// TIA Portal project "CurrentConfig" (V16)

(* hardware
DEVICE "ET 200S station_1"  ET 200S station
   slot 0: "Rack"  Rail
   slot 2: "-20K0 - PLC"  IM151-8 PN/DP CPU  6ES7 151-8AB01-0AB0  V3.2
      slot 1: "PROFINET interface_1"  PN-IO
         slot 1: "Port_1"  Port
         slot 2: "Port_2"  Port
         slot 3: "Port_3"  Port
   slot 4: "-20K1 - VOEDING"  PM-E 24VDC  6ES7 138-4CA01-0AA0
   slot 5: "-20K2 - INGANG_1"  8DI DC24V  6ES7 131-4BF00-0AA0
   slot 6: "-20K3 - INGANG_2"  8DI DC24V  6ES7 131-4BF00-0AA0
   slot 7: "-20K4 - INGANG_3"  8DI DC24V  6ES7 131-4BF00-0AA0
   slot 8: "-20K5 - INGANG_4"  8DI x 24VDC  6ES7 131-4BF00-0AA0
   slot 9: "-20K6 - UITGANG_1"  8DO x 24VDC / 0.5A  6ES7 132-4BF00-0AA0
   slot 10: "8DO x 24VDC / 0.5A_1"  8DO x 24VDC / 0.5A  6ES7 132-4BF00-0AA0
   slot 11: "PM-E 24VDC_1"  PM-E 24VDC  6ES7 138-4CA01-0AA0
   slot 12: "-20K8 - UITGANG_2"  8DO x 24VDC / 0.5A  6ES7 132-4BF00-0AA0
   slot 13: "-20K9 - UITGANG_3"  8DO x 24VDC / 0.5A  6ES7 132-4BF00-0AA0
   slot 14: "-20K10 - UITGANG_4"  8DO x 24VDC / 0.5A  6ES7 132-4BF00-0AA0
   slot 15: "-20K11 - UITGANG_5"  8DO x 24VDC / 0.5A  6ES7 132-4BF00-0AA0
   slot 16: "-20K12 - UITGANG_6 (4)"  4DO x 24VDC / 0.5A ST  6ES7 132-4BD02-0AA0
   slot 17: "-20K13 - UITGANG_7 (4)"  4DO x 24VDC / 0.5A ST  6ES7 132-4BD02-0AA0
   slot 18: "1 Count 24V Encoder Wals"  1 COUNT 24V  6ES7 138-4DA04-0AB0  V2.0
   slot 19: "1 Count 24V Encoder Band"  1 COUNT 24V  6ES7 138-4DA04-0AB0  V2.0
DEVICE "HMI_1"  KTP700 Basic PN
   slot 0: "HMI_1"  KTP700 Basic PN  6AV2 123-2GB03-0AX0  16.0.0.0
   slot 1: "HMI_RT_2"  KTP700 Basic PN  6AV2 123-2GB03-0AX0  16.0.0.0
   slot 5: "HMI_1.IE_CP_1"  PROFINET Interface  16.0.0.0
      slot 1: "PROFINET Interface_1"  PROFINET Interface
         slot 1: "Port_1"  Port
*)

// ===== PLC "-20K0 - PLC"  IM151-8 PN/DP CPU =====

VAR_GLOBAL   // PLC tag table "Default tag table"
   "Drive 1 Ready" AT %I0.0 : Bool;   // +MC-21K2:1 - Drive 1 Ready
   "Drive 2 Ready" AT %I0.1 : Bool;   // +MC-21K2:5 - Drive 2 Ready
   "Drive 3 Ready" AT %I0.2 : Bool;   // +MC-21K2:2 - Drive 3 Ready
   "Drive 4 Ready" AT %I0.3 : Bool;   // +MC-21K2:6 - Drive 4 Ready
   "Drive 5 Ready" AT %I0.4 : Bool;   // +MC-21K2:3 - Drive 5 Ready
   "Sensor Trechter" AT %I0.5 : Bool;   // +MC-21K2:7 - Sensor Trechter
   "Sensor Op Band" AT %I0.6 : Bool;   // +MC-21K2:4 Sensor Op Band
   "Sensor Wals (Option)" AT %I0.7 : Bool;   // +MC-21K2:8 - Sensor Wals (Option)
   "ESB Oke" AT %I1.0 : Bool;   // +MC-21K3:1 - ESB Oke
   "ESB Pressend" AT %I1.1 : Bool;   // +MC-21K3:5 - ESB Pressend
   "Reset Active" AT %I1.2 : Bool;   // +MC-21K3:2 - Reset Active
   "Noodsleutel(1)" AT %I1.3 : Bool;   // +MC-21K3:6 - NOODSLEUTEL
   "Alle uitgangen(1)" AT %I1.4 : Bool;   // +MC-21K3:3 - Alle uitgangen
   "Door 1 NC contact" AT %I1.5 : Bool;   // +MC-21K3:7 - Safety Doorswitch 1
   "Door 1 NO contact" AT %I1.6 : Bool;   // +MC-21K3:4 - Safety Doorswitch 1 Normaly open
   "Door 2 NC contact" AT %I1.7 : Bool;   // +MC-21K3:8 - Safety Doorswitch 2
   "Spare(5)" AT %I3.0 : Bool;
   "Spare(6)" AT %I3.1 : Bool;
   "Spare(10)" AT %I180.0 : Bool;   // Spare
   "Spare(11)" AT %I180.1 : Bool;   // Spare
   "Spare(12)" AT %I3.4 : Bool;   // Spare
   "Spare(13)" AT %I3.5 : Bool;   // Spare
   "Spare(14)" AT %I3.6 : Bool;   // Spare
   "Spare(15)" AT %I3.7 : Bool;   // Spare
   "Programma 1" AT %I2.0 : Bool;   // +MC-21K4:1 - Programma 1
   "Programma 2" AT %I2.1 : Bool;   // +MC-21K4:5 - Programma 2 (Option)
   "Programma 3" AT %I2.2 : Bool;   // +MC-21K4:2 - Programma 3
   "Cleaning" AT %I2.3 : Bool;   // +MC-21K4:6 - Cleaning
   "Start Machine" AT %I2.4 : Bool;   // +MC-21K4:3 - Start Machine
   "Stop Machine" AT %I2.5 : Bool;   // +MC-21K4:7 - Stop Machine
   "Spare(16)" AT %I2.6 : Bool;   // Spare
   "Encoder_Z_Puls" AT %I2.7 : Bool;   // Spare
   "Safety Relais" AT %Q0.0 : Bool;   // +MC-21K6:1 - Safety Relais
   "Bel Storing" AT %Q0.1 : Bool;   // +MC-21K6:5 - Bel Storing
   "Spare" AT %Q5.3 : Bool;   // Spare
   "Drive 1 RUN FWD" AT %Q1.0 : Bool;   // +MC-21K8:1 - Drive 1 RUN FWD
   "Drive 1 REV]" AT %Q1.1 : Bool;   // +MC-21K8:5 - Drive 1 REV
   "Drive 1 Speed 1" AT %Q1.2 : Bool;   // +MC-21K8:2 - Drive 1 Speed 1
   "Drive 1 Speed 2" AT %Q1.3 : Bool;   // +MC-21K8:6 - Drive 1 Speed 2
   "Spare(3)" AT %Q1.4 : Bool;   // Spare
   "Drive 2 RUN FWD" AT %Q1.5 : Bool;   // +MC-21K8:7 - Drive 2 RUN FWD
   "Drive 2 REV" AT %Q1.6 : Bool;   // +MC-21K8:4 - Drive 2 REV
   "Drive 2 Speed 1" AT %Q1.7 : Bool;   // +MC-21K8:8 - Drive 2 Speed 1
   "Drive 2 Speed 2" AT %Q2.0 : Bool;   // +MC-21K9:1 - Drive 2 Speed 2
   "Spare(4)" AT %Q2.1 : Bool;   // Spare
   "Drive 3 RUN FWD" AT %Q2.2 : Bool;   // +MC-21K9:2 - Drive 3 RUN FWD
   "Drive 3 REV" AT %Q2.3 : Bool;   // +MC-21K9:6 - Drive 3 REV
   "Drive 3 Speed 1" AT %Q2.4 : Bool;   // +MC-21K9:3 - Drive 3 Speed 1
   "Drive 3 Speed 2" AT %Q2.5 : Bool;   // +MC-21K9:7 - Drive 3 Speed 2
   "Spare(21)" AT %Q2.6 : Bool;   // Spare
   "Drive 4 RUN FWD" AT %Q2.7 : Bool;   // +MC-21K9:8 - Drive 4 RUN FWD
   "Drive 4 REV" AT %Q3.0 : Bool;   // +MC-21K10:1 - Drive 4 REV
   "Drive 4 Speed 1" AT %Q3.1 : Bool;   // +MC-21K10:5 - Drive 4 Speed 1
   "Drive 4 Speed 2" AT %Q3.2 : Bool;   // +MC-21K10:2 - Drive 4 Speed 2
   "Spare(22)" AT %Q3.3 : Bool;   // Spare
   "Drive 5 RUN FWD" AT %Q3.4 : Bool;   // +MC-21K10:3 - Drive 5 RUN FWD
   "Drive 5 REV" AT %Q3.5 : Bool;   // +MC-21K10:7 - Drive 5 REV
   "Drive 5 Speed 1" AT %Q3.6 : Bool;   // +MC-21K10:4 - Drive 5 Speed 1
   "Drive 5 Speed 2" AT %Q3.7 : Bool;   // +MC-21K10:8 - Drive 5 Speed 2
   "Spare(23)" AT %Q4.0 : Bool;   // Spare
   "LED Programma 1" AT %Q4.1 : Bool;   // +MC-21K11:5 - LED Programma 1
   "LED Programma 2" AT %Q4.2 : Bool;   // +MC-21K11:2 - LED Programma 2
   "LED Programma 3" AT %Q4.3 : Bool;   // +MC-21K11:6 - LED Programma 3
   "LED E-STOP" AT %Q0.2 : Bool;   // +MC-21K6:2- LED E-STOP
   "LED RUN" AT %Q4.5 : Bool;   // +MC-21K11:7 - LED RUN
   "Valve 1" AT %Q4.6 : Bool;   // +MC-21K11:4 - Valve 1
   "Valve 2" AT %Q4.7 : Bool;   // +MC-21K11:8 - Valve 2
   "Valve 3" AT %Q5.0 : Bool;   // +MC-21K12:1 - Valve 3
   "Valve 4" AT %Q5.1 : Bool;   // +MC-21K12:5 - Valve 4
   "Valve 5" AT %Q5.2 : Bool;   // +MC-21K12:2 - Valve 5
   "Spare(1)" AT %Q6.0 : Bool;   // Spare
   "Spare(2)" AT %Q6.1 : Bool;   // Spare
   "Spare(18)" AT %Q6.2 : Bool;   // Spare
   "Spare(19)" AT %Q6.3 : Bool;   // Spare
   "Spare(20)" AT %Q4.4 : Bool;   // Spare
   "Drive 1 Rapid Stop" AT %Q0.3 : Bool;   // +MC-21K6:6 - Drive 1 Rapid Stop
   "Drive 2 Rapid Stop" AT %Q0.4 : Bool;   // +MC-21K6:3 - Drive 2 Rapid Stop
   "Drive 3 Rapid Stop" AT %Q0.5 : Bool;   // +MC-21K6:7 - Drive 3 Rapid Stop
   "Drive 4 Rapid Stop" AT %Q0.6 : Bool;   // +MC-21K6:4 - Drive 4 Rapid Stop
   "Drive 5 Rapid Stop" AT %Q0.7 : Bool;   // +MC-21K6:8 - Drive 5 Rapid Stop
   "Systeem RUN" AT %M0.0 : Bool;   // Systeem RUN
   "Tag_1" AT %M0.1 : Bool;
   "Tag_2" AT %M0.2 : Bool;
   "Tag_3" AT %M0.3 : Bool;
   "Tag_4" AT %M0.4 : Bool;
   "Safety Feedback" AT %M0.6 : Bool;
   "Tag_5" AT %M0.7 : Bool;
   "Tag_6" AT %M1.0 : Bool;
   "ONC Drive 1 RUN FWD" AT %M10.0 : Bool;
   "ONC Drive 2 RUN FWD" AT %M10.1 : Bool;
   "ONC Drive 3 RUN FWD" AT %M10.2 : Bool;
   "ONC Drive 4 RUN FWD" AT %M10.3 : Bool;
   "ONC Drive 5 RUN FWD" AT %M10.4 : Bool;
   "ONC Drive 1 RUN FWD and Speed 1" AT %M10.5 : Bool;
   "ONC Drive 2 RUN FWD and Speed 1" AT %M10.6 : Bool;
   "ONC Drive 3 RUN FWD and Speed 1" AT %M10.7 : Bool;
   "ONC Drive 4 RUN FWD and Speed 1" AT %M11.0 : Bool;
   "ONC Drive 5 RUN FWD and Speed 1" AT %M11.1 : Bool;
   "ONC Drive 1 RUN FWD and Speed 2" AT %M11.2 : Bool;
   "ONC Drive 2 RUN FWD and Speed 2" AT %M11.3 : Bool;
   "ONC Drive 3 RUN FWD and Speed 2" AT %M11.4 : Bool;
   "ONC Drive 4 RUN FWD and Speed 2" AT %M11.5 : Bool;
   "ONC Drive 5 RUN FWD and Speed 2" AT %M11.6 : Bool;
   "Startknop_Scherm" AT %M15.0 : Bool;
   "Stopknop_Scherm" AT %M15.1 : Bool;
   "Tag_7" AT %M110.1 : Bool;
   "Reset_scherm" AT %M15.2 : Bool;
   "Sensor_op_band_memory" AT %M15.3 : Bool;
   "System RUN_1" AT %M20.0 : Bool;
   "ResetDelay" AT %M20.1 : Bool;
   "SensorWalsMemory" AT %M20.2 : Bool;
   "Timer_Memory" AT %M20.3 : Bool;
   "StopAll" AT %M20.4 : Bool;
   "Tag_8" AT %M100.3 : Bool;
   "Tag_9" AT %M100.4 : Bool;
   "Tag_10" AT %M0.5 : Bool;
   "Tag_11" AT %M150.0 : Bool;
   "Tag_12" AT %M101.1 : Bool;
   "Tag_13" AT %T1 : Timer;
   "Tag_14" AT %M300.0 : Bool;
   "Tag_15" AT %M260.0 : Bool;
   "Tag_16" AT %M300.1 : Bool;
   "Tag_17" AT %M501.0 : Bool;
   "Tag_18" AT %M500.1 : Bool;
   "Tag_19" AT %M160.0 : Bool;
   "Tag_20" AT %M150.5 : Bool;
   "Tag_21" AT %QD256 : DWord;
   "Tag_22" AT %QW260 : Word;
   "Tag_23" AT %ID256 : DWord;
   "Tag_24" AT %ID260 : DWord;
   "Tag_25" AT %ID464 : DWord;
   "Tag_26" AT %ID471 : DWord;
   "Tag_27" AT %QW471 : Word;
   "Tag_28" AT %QD464 : DWord;
   "Tag_30" AT %IW205 : Int;
   "SystemTime" AT %MD2 : Time;
   "Tag_31" AT %M5.0 : Bool;
   "Lamp_Green" AT %Q7.0 : Bool;
   "Lamp_Blue" AT %Q7.1 : Bool;
   "Lamp_Yellow" AT %Q7.2 : Bool;
   "Lamp_Red" AT %Q7.3 : Bool;
   "Lamp_Buzzer" AT %Q7.4 : Bool;
   "PulseTimer" AT %T0 : Timer;
END_VAR

VAR_GLOBAL   // PLC tag table "Outputs/HMI"
   "Drive_1_Auto" AT %M50.0 : Bool;
   "Drive_1_Manual" AT %M50.1 : Bool;
   "Drive_2_Auto" AT %M50.2 : Bool;
   "Drive_2_Manual" AT %M50.3 : Bool;
   "Drive_3_Auto" AT %M50.4 : Bool;
   "Drive_3_Manual" AT %M50.5 : Bool;
   "Drive_4_Auto" AT %M50.6 : Bool;
   "Drive_4_Manual" AT %M50.7 : Bool;
   "Drive_5_Auto" AT %M51.0 : Bool;
   "Drive_5_Manual" AT %M51.1 : Bool;
   "Valve_1_Auto" AT %M51.2 : Bool;
   "Valve_1_Manual" AT %M51.3 : Bool;
   "Valve_2_Auto" AT %M51.4 : Bool;
   "Valve_2_Manual" AT %M51.5 : Bool;
   "Valve_3_Auto" AT %M51.6 : Bool;
   "Valve_3_Manual" AT %M51.7 : Bool;
   "Valve_4_Auto" AT %M52.0 : Bool;
   "Valve_4_Manual" AT %M52.1 : Bool;
   "Valve_5_Auto" AT %M52.2 : Bool;
   "Valve_5_Manual" AT %M52.3 : Bool;
   "Stop_drive_1" AT %M52.4 : Bool;
   "Stop_drive_2" AT %M52.5 : Bool;
   "Stop_drive_3" AT %M52.6 : Bool;
   "Stop_drive_4" AT %M52.7 : Bool;
   "Stop_drive_5" AT %M53.0 : Bool;
   "Stop_valve_1" AT %M53.1 : Bool;
   "Stop_valve_2" AT %M53.2 : Bool;
   "Stop_valve_3" AT %M53.3 : Bool;
   "Stop_valve_4" AT %M53.4 : Bool;
   "Stop_valve_5" AT %M53.5 : Bool;
   "Trechter_Bijvullen_Signaal" AT %M53.6 : Bool;
   "LED_ESB01" AT %M53.7 : Bool;
   "LED_MagazijnStoring" AT %M54.0 : Bool;
   "Alarm_Axis_Not_Position" AT %M54.1 : Bool;
   "Alarm_Product_Not_Position" AT %M54.2 : Bool;
   "Door_Safety_Alarm" AT %M54.3 : Bool;
   "ESB_Safety_Alarm" AT %M54.4 : Bool;
   "Alarms(1)" AT %MW500 : Word;
   "HMI_Des_Pos_Axis3" AT %M54.5 : Bool;
   "GoButtonPressed" AT %M54.6 : Bool;
   "Drive_3_ReferencePos" AT %M54.7 : Bool;
   "SequenceStep" AT %MW55 : Int;
   "Drive_3_ReferencePos_Active" AT %M58.0 : Bool;
   "Start_Axis3_Procedure" AT %M58.1 : Bool;
   "ProductProcessed" AT %M58.2 : Bool;
   "GoToNextProduct" AT %M60.0 : Bool;
   "Product_Counter" AT %MW58 : Int;
   "Axis_3_On_RefPos" AT %M62.0 : Bool;
   "TimerProductRAM" AT %MW57 : Int;
   "TimerCounterValue" AT %MW64 : Int;
   "Prev_Sensor_Op_Band" AT %M180.0 : Bool;
   "CurrentCycle" AT %MW180 : Int;
   "Naar_Pos_0" AT %M180.1 : Bool;
   "Cleaning_Active" AT %M182.0 : Bool;
   "Cleaning_Confirmed" AT %M182.1 : Bool;
   "Cleaning_Cancelled" AT %M182.2 : Bool;
   "Cleaning_Screen_Active" AT %M182.3 : Bool;
   "CleaningEnd" AT %M182.4 : Bool;
   "HMI_ManualControl" AT %M182.5 : Bool;
   "Drive_3_Manual_Rev" AT %M60.1 : Bool;
   "Drive_3_FastStop" AT %M60.2 : Bool;
END_VAR

VAR_GLOBAL   // PLC tag table "Secund. Tags"
   "Aanvoerband_Tag1" AT %M100.0 : Bool;
   "Aanvoerband_Tag2" AT %M100.1 : Bool;
   "Trechter_Bijvullen_Haltveroorzaker" AT %M100.2 : Bool;
   "Safety_Automatic" AT %M100.5 : Bool;
   "Safety_Override" AT %M100.6 : Bool;
   "RUN_Automatic" AT %M100.7 : Bool;
   "RUN_Manual" AT %M101.0 : Bool;
   "Invert_Trechter_Sensor" AT %M101.2 : Bool;
   "WalsSensorMemory" AT %M101.3 : Bool;
   "Disable_Module" AT %M101.4 : Bool;
   "Sensor_Trechter_Delayed" AT %M101.5 : Bool;
   "Positive_Flank" AT %M101.6 : Bool;
   "ProductSensor_Flank" AT %M101.7 : Bool;
   "ProductSensor_Rug" AT %M102.0 : Bool;
   "SensorRug" AT %M102.1 : Bool;
   "TimeCyclusEnd" AT %M102.2 : Bool;
   "CounterReset" AT %M102.3 : Bool;
   "StartTimer" AT %M102.4 : Bool;
   "StopTimer" AT %M102.5 : Bool;
   "SaveTimervalue" AT %M102.6 : Bool;
   "ResetTotalProducts" AT %M102.7 : Bool;
   "MaintenanceNeeded" AT %M103.0 : Bool;
   "RetainValues" AT %M112.0 : Bool;
   "Retain_1_DontTouch!" AT %M112.1 : Bool;
   "Safety_Doors" AT %M112.2 : Bool;
   "Overname_Linked_Drive1" AT %M112.3 : Bool;
   "Drive_RefuseLinkingDrive1" AT %M112.4 : Bool;
   "Drive_4_Speed1_Link" AT %M112.5 : Bool;
   "Drive_4_Speed1_Unlink" AT %M112.6 : Bool;
   "SafetyOK" AT %M112.7 : Bool;
   "Valve2_Pulse" AT %M113.0 : Bool;
END_VAR

VAR_GLOBAL   // PLC tag table "PositionControl"
   "Counter1_IW100" AT %IW100 : Int;
   "Counter2_IW102" AT %IW102 : Int;
   "Manual Jog Fwd" AT %M137.0 : Bool;
   "Manual Jog Rev" AT %M137.1 : Bool;
   "ReferenceSwitchAxis3" AT %I3.0 : Bool;
   "EncoderBand_Alive" AT %IW110 : Int;
   "EncoderBand_RawCounter" AT %IW112 : Int;
   "EncoderBand_FineCounter" AT %IW113 : Int;
   "Zpuls_Encoder_Band" AT %I110.3 : Bool;
END_VAR

TYPE "ProductEntry"
   STRUCT
      StartTime : Time := T#0ms;
      Active : Bool;
   END_STRUCT;
END_TYPE

TYPE "ProductTrack"
   STRUCT
      StartPosition : Real;
      Active : Bool;
   END_STRUCT;
END_TYPE

DATA_BLOCK "ProductBuffer_V3_DB"   // DB90
{ S7_Optimized_Access := 'FALSE' }
VERSION : 0.1
// stored: InstanceOfName ProductBuffer_V3
"ProductBuffer_V3"
BEGIN
END_DATA_BLOCK

// folder: 1000 Data

DATA_BLOCK "PLCMemory"   // DB15
{ S7_Optimized_Access := 'FALSE' }
VERSION : 0.1
   VAR
      Homing_Sensor_Wals_Offset_Test : Time := T#1S_200MS;   // Offset of homing position sensor wals
      Wals_Delay_Offset : Time := T#400MS;   // Offset of Wals on delay
      Safety_Delay : Time := T#5MS;   // Delay of safety high
      WalsCheck_Time : Time := T#5S;   // Time offset when wals slipping message is displayed
      ProductCheck_Time : Time := T#15S;   // Time offset when aanvoer not in position message is displayed
      ProductIntervalTime : Time;   // Counts the time between 2 products
      ProductIntervalTime_1 : Time;   // Depends on ProductIntervalTimer
      ProductIntervalTime_2 : Time;   // Depends on ProductIntervalTimer_1
      TD_Products_Counter : Int;   // Counts the total amount of products with the Sensor Band
      UsernameMemory : String := 'Key';
      PasswordMemory : String := 'Key123';
      SpeedSettingsTakeover : Bool := True;   // Makes the speed of Overname the same as speed Drive 1
      SpeedSettingOvername : Bool;   // Parameter of setting the speed for Drive 4 (Overname)
      SpeedSettingBand : Bool;   // Parameter of setting the speed for Drive 1 (Band)
      TimingSettingOvername : Bool := True;   // Makes the timing of Overname the same as speed Drive 1
      EncoderPosition : Real;   // Real Value of Encoder Axis 3 (Wals)
      StepSize : Real := 0.0;   // Pulsfactor of Encoder Axis 3
      Desired_Encoder_Position : Real;
      Tolerance : Real := 0.0;
      "Encoder PulsOffset" : Time := T#3MS;
      Axis3_Ref_Pos : Real := 85.0;   // Refention position of Axis 3 without tolerance
      Reference_Position_Axis3 : Real;   // Refention position of Axis 3 with calculated tolerance
      ProductCount : Int;
      Axis3_ControlMode : Bool := true;
      Axis1_ControlMode : Bool := true;
      ProductsToProduce : Int;
      SystemTime : Time;
      Disable_Modules : Struct
         Disable_Band : Bool;
         Disable_Trilgoten : Bool;
         Disable_AanvoerWals : Bool;
         Disable_Aandruk1 : Bool;
         Disable_Aandruk2 : Bool;
         Disable_Aandruk3 : Bool;
         Disable_Blaaspuls : Bool;
         Disable_Retourband : Bool;
         Disable_Afsluiter : Bool;
      END_STRUCT;
      Offset_Timers : Struct
         Trilgoten_Start_Offset : Time := T#10MS;   // Delay offset of start trilgoten
         Trilgoten_Stop_Offset : Time := T#10MS;   // Delay offset of stop trilgoten
         Aanvoer_Start_Offset : Time := T#10MS;   // Delay offset of start aanvoer
         Magazijn_Sensor_Delay : Time := T#15S;   // Delay on magazijn sensor.
         Aanvoer_Stop_Offset : Time := T#10MS;   // Delay offset of stop aanvoer
         Overname_Start_Offset : Time := T#5MS;   // Delay offset of start Overname
         Overname_Stop_Offset : Time := T#5MS;   // Delay offset of stop Overname
         Retourband_Start_Offset : Time := T#5ms;
         Retourband_Stop_Offset : Time := T#5ms;
         BlowOff_CycleTime : Time := T#500ms;
         Blow_Off_PulseTime : Time := T#500ms;
      END_STRUCT;
      ProductBuffer : Struct
         DelayTime : Time := T#7s;
         ProductsCount : Int;
         MoveTrigger : Bool;
         MoveFeedback : Bool;
         RestFeedback : Bool;
         InsertIndex : Int;
      END_STRUCT;
      ProductBufferBehindWals : Struct
         DelayTime : Time := T#2s_500MS;
         Product_Count : Int;
      END_STRUCT;
   END_VAR
BEGIN
END_DATA_BLOCK

DATA_BLOCK "FB_SystemTimeCounter_DB_1"   // DB23
{ S7_Optimized_Access := 'FALSE' }
VERSION : 0.1
// stored: InstanceOfName FB_SystemTimeCounter
"FB_SystemTimeCounter"
BEGIN
END_DATA_BLOCK

DATA_BLOCK "ResetOuputs_Function_Rest"   // DB29
{ S7_Optimized_Access := 'FALSE' }
VERSION : 0.1
// stored: InstanceOfName ResetOuputs_Function
"ResetOuputs_Function"
BEGIN
END_DATA_BLOCK

DATA_BLOCK "ProductBuffer_DB"   // DB58
{ S7_Optimized_Access := 'FALSE' }
VERSION : 0.1
// stored: InstanceOfName ProductBuffer
"ProductBuffer"
BEGIN
END_DATA_BLOCK

DATA_BLOCK "MC_Move_Prog.1_1"   // DB59
{ S7_Optimized_Access := 'FALSE' }
VERSION : 0.1
// stored: InstanceOfName MC_Move
"MC_Move"
BEGIN
END_DATA_BLOCK

DATA_BLOCK "MC_Move_DB"   // DB62
{ S7_Optimized_Access := 'FALSE' }
VERSION : 0.1
// stored: InstanceOfName MC_Move
"MC_Move"
BEGIN
END_DATA_BLOCK

DATA_BLOCK "Blinker_BlueBlinking"   // DB63
{ S7_Optimized_Access := 'FALSE' }
VERSION : 0.1
// stored: InstanceOfName Blinker
"Blinker"
BEGIN
END_DATA_BLOCK

DATA_BLOCK "Programma 1 - Test_DB"   // DB64
{ S7_Optimized_Access := 'FALSE' }
VERSION : 0.1
// stored: InstanceOfName Programma 1 - Test
"Programma 1 - Test"
BEGIN
END_DATA_BLOCK

DATA_BLOCK "Blinker_BlueConstant"   // DB65
{ S7_Optimized_Access := 'FALSE' }
VERSION : 0.1
// stored: InstanceOfName Blinker
"Blinker"
BEGIN
END_DATA_BLOCK

DATA_BLOCK "ProductBuffer_V2_DB"   // DB66
{ S7_Optimized_Access := 'FALSE' }
VERSION : 0.1
// stored: InstanceOfName ProductBuffer_V2
"ProductBuffer_V2"
BEGIN
END_DATA_BLOCK

DATA_BLOCK "FB_ProductTrigger_1"   // DB67
{ S7_Optimized_Access := 'FALSE' }
VERSION : 0.1
// stored: InstanceOfName FB_ProductTrigger
"FB_ProductTrigger"
BEGIN
END_DATA_BLOCK

DATA_BLOCK "BlowOff_Timer_Cleaning"   // DB73
{ S7_Optimized_Access := 'FALSE' }
VERSION : 0.1
// stored: InstanceOfName BlowOff_Timer
"BlowOff_Timer"
BEGIN
END_DATA_BLOCK

DATA_BLOCK "Blinker_BlowOff"   // DB74
{ S7_Optimized_Access := 'FALSE' }
VERSION : 0.1
// stored: InstanceOfName Blinker
"Blinker"
BEGIN
END_DATA_BLOCK

DATA_BLOCK "BlowOff_Timer_Prog1"   // DB75
{ S7_Optimized_Access := 'FALSE' }
VERSION : 0.1
// stored: InstanceOfName BlowOff_Timer
"BlowOff_Timer"
BEGIN
END_DATA_BLOCK

DATA_BLOCK "MC_Move_1"   // DB76
{ S7_Optimized_Access := 'FALSE' }
VERSION : 0.1
// stored: InstanceOfName MC_Move
"MC_Move"
BEGIN
END_DATA_BLOCK

DATA_BLOCK "MC_Move_2"   // DB77
{ S7_Optimized_Access := 'FALSE' }
VERSION : 0.1
// stored: InstanceOfName MC_Move
"MC_Move"
BEGIN
END_DATA_BLOCK

DATA_BLOCK "FB_EncoderFeedback_Aanvoerband"   // DB78
{ S7_Optimized_Access := 'FALSE' }
VERSION : 0.1
// stored: InstanceOfName FB_EncoderFeedback_Degree
"FB_EncoderFeedback_Degree"
BEGIN
END_DATA_BLOCK

DATA_BLOCK "ProductBuffer_BehindWals"   // DB79
{ S7_Optimized_Access := 'FALSE' }
VERSION : 0.1
// stored: InstanceOfName ProductBuffer
"ProductBuffer"
BEGIN
END_DATA_BLOCK

DATA_BLOCK "Blinker_GreenConstant"   // DB81
{ S7_Optimized_Access := 'FALSE' }
VERSION : 0.1
// stored: InstanceOfName Blinker
"Blinker"
BEGIN
END_DATA_BLOCK

DATA_BLOCK "ProductBuffer_V2_DB_BehindWals"   // DB82
{ S7_Optimized_Access := 'FALSE' }
VERSION : 0.1
// stored: InstanceOfName ProductBuffer_V2
"ProductBuffer_V2"
BEGIN
END_DATA_BLOCK

DATA_BLOCK "BlowOff_Timer_ManualDB"   // DB83
{ S7_Optimized_Access := 'FALSE' }
VERSION : 0.1
// stored: InstanceOfName BlowOff_Timer
"BlowOff_Timer"
BEGIN
END_DATA_BLOCK

DATA_BLOCK "ProductBuffer_DB_Manual"   // DB85
{ S7_Optimized_Access := 'FALSE' }
VERSION : 0.1
// stored: InstanceOfName ProductBuffer
"ProductBuffer"
BEGIN
END_DATA_BLOCK

DATA_BLOCK "BlowOff_Timer_Manual2DB"   // DB86
{ S7_Optimized_Access := 'FALSE' }
VERSION : 0.1
// stored: InstanceOfName BlowOff_Timer
"BlowOff_Timer"
BEGIN
END_DATA_BLOCK

// folder: 900 Systeem

DATA_BLOCK "DB_SystemTimeCounter"   // DB68
{ S7_Optimized_Access := 'FALSE' }
VERSION : 0.1
   VAR
      SystemTime : Time;
   END_VAR
BEGIN
END_DATA_BLOCK

DATA_BLOCK "FB_SystemTimeCounter_DB"   // DB69
{ S7_Optimized_Access := 'FALSE' }
VERSION : 0.1
// stored: InstanceOfName FB_SystemTimeCounter
"FB_SystemTimeCounter"
BEGIN
END_DATA_BLOCK

// folder: Blocks

DATA_BLOCK "SwitchBlockAxisPosition_DB"   // DB39
{ S7_Optimized_Access := 'FALSE' }
VERSION : 0.1
// stored: InstanceOfName SwitchBlockAxisPosition
"SwitchBlockAxisPosition"
BEGIN
END_DATA_BLOCK

DATA_BLOCK "Blinker_Start"   // DB71
{ S7_Optimized_Access := 'FALSE' }
VERSION : 0.1
// stored: InstanceOfName Blinker
"Blinker"
BEGIN
END_DATA_BLOCK

// folder: Functions

DATA_BLOCK "2in-1out_Block_LED-Estop"   // DB1
{ S7_Optimized_Access := 'FALSE' }
VERSION : 0.1
// stored: InstanceOfName 2in-1out_Block
"2in-1out_Block"
BEGIN
END_DATA_BLOCK

DATA_BLOCK "2in-1out_Block_Start/Stop_Override"   // DB2
{ S7_Optimized_Access := 'FALSE' }
VERSION : 0.1
// stored: InstanceOfName 2in-1out_Block
"2in-1out_Block"
BEGIN
END_DATA_BLOCK

DATA_BLOCK "Override_Block_Safety_1"   // DB3
{ S7_Optimized_Access := 'FALSE' }
VERSION : 0.1
// stored: InstanceOfName Override_Block_Safety
"Override_Block_Safety"
BEGIN
END_DATA_BLOCK

DATA_BLOCK "Ouput_Function_1_Drive1"   // DB4
{ S7_Optimized_Access := 'FALSE' }
VERSION : 0.1
// stored: InstanceOfName Ouput_Function_1
"Ouput_Function_1"
BEGIN
END_DATA_BLOCK

DATA_BLOCK "Ouput_Function_1_Drive2"   // DB8
{ S7_Optimized_Access := 'FALSE' }
VERSION : 0.1
// stored: InstanceOfName Ouput_Function_1
"Ouput_Function_1"
BEGIN
END_DATA_BLOCK

DATA_BLOCK "Ouput_Function_1_Drive3"   // DB12
{ S7_Optimized_Access := 'FALSE' }
VERSION : 0.1
// stored: InstanceOfName Ouput_Function_1
"Ouput_Function_1"
BEGIN
END_DATA_BLOCK

DATA_BLOCK "Ouput_Function_1_Drive4"   // DB17
{ S7_Optimized_Access := 'FALSE' }
VERSION : 0.1
// stored: InstanceOfName Ouput_Function_1
"Ouput_Function_1"
BEGIN
END_DATA_BLOCK

DATA_BLOCK "Ouput_Function_1_Drive5"   // DB18
{ S7_Optimized_Access := 'FALSE' }
VERSION : 0.1
// stored: InstanceOfName Ouput_Function_1
"Ouput_Function_1"
BEGIN
END_DATA_BLOCK

DATA_BLOCK "Ouput_Function_1_Valve1"   // DB19
{ S7_Optimized_Access := 'FALSE' }
VERSION : 0.1
// stored: InstanceOfName Ouput_Function_1
"Ouput_Function_1"
BEGIN
END_DATA_BLOCK

DATA_BLOCK "Alarms"   // DB24
{ S7_Optimized_Access := 'FALSE' }
VERSION : 0.1
   VAR
      AlarmStruct : Struct
         Alarm_Product_Not_Position : Bool;
         Alarm_Axis_Not_Position : Bool;
         Alarm_Drive1 : Bool;
         Alarm_Drive2 : Bool;
         Alarm_Drive3 : Bool;
         Alarm_Drive4 : Bool;
         Alarm_Drive5 : Bool;
         "Alarm_To_Many_Products_Reset_Counter!" : Bool;
      END_STRUCT;
      AlarmsWord : Word;
      HMI_Alarm_Drive1 : Word;
      HMI_Alarm_Drive2 : Word;
      HMI_Alarm_Drive3 : Word;
      HMI_Alarm_Drive4 : Word;
      HMI_Alarm_Drive5 : Word;
   END_VAR
BEGIN
END_DATA_BLOCK

DATA_BLOCK "Ouput_Function_1_Valve2"   // DB25
{ S7_Optimized_Access := 'FALSE' }
VERSION : 0.1
// stored: InstanceOfName Ouput_Function_1
"Ouput_Function_1"
BEGIN
END_DATA_BLOCK

DATA_BLOCK "Ouput_Function_1_Valve3"   // DB26
{ S7_Optimized_Access := 'FALSE' }
VERSION : 0.1
// stored: InstanceOfName Ouput_Function_1
"Ouput_Function_1"
BEGIN
END_DATA_BLOCK

DATA_BLOCK "Ouput_Function_1_Valve4"   // DB27
{ S7_Optimized_Access := 'FALSE' }
VERSION : 0.1
// stored: InstanceOfName Ouput_Function_1
"Ouput_Function_1"
BEGIN
END_DATA_BLOCK

DATA_BLOCK "Ouput_Function_1_Valve5"   // DB28
{ S7_Optimized_Access := 'FALSE' }
VERSION : 0.1
// stored: InstanceOfName Ouput_Function_1
"Ouput_Function_1"
BEGIN
END_DATA_BLOCK

DATA_BLOCK "ESB_Buzzer_Block"   // DB33
{ S7_Optimized_Access := 'FALSE' }
VERSION : 0.1
// stored: InstanceOfName ESB_Flash_Warning_Block
"ESB_Flash_Warning_Block"
BEGIN
END_DATA_BLOCK

DATA_BLOCK "ESB_Lamp_Block"   // DB34
{ S7_Optimized_Access := 'FALSE' }
VERSION : 0.1
// stored: InstanceOfName ESB_Flash_Warning_Block
"ESB_Flash_Warning_Block"
BEGIN
END_DATA_BLOCK

DATA_BLOCK "Delayed_Message_Function_Magazine"   // DB38
{ S7_Optimized_Access := 'FALSE' }
VERSION : 0.1
// stored: InstanceOfName Delayed_Message_Function
"Delayed_Message_Function"
BEGIN
END_DATA_BLOCK

DATA_BLOCK "Alarm_Axis_Position_Function_Wals"   // DB41
{ S7_Optimized_Access := 'FALSE' }
VERSION : 0.1
// stored: InstanceOfName Alarm_Axis_Position_Function
"Alarm_Axis_Position_Function"
BEGIN
END_DATA_BLOCK

DATA_BLOCK "Alarm_Axis_Position_Function_Wals1"   // DB42
{ S7_Optimized_Access := 'FALSE' }
VERSION : 0.1
// stored: InstanceOfName Alarm_Axis_Position_Function
"Alarm_Axis_Position_Function"
BEGIN
END_DATA_BLOCK

DATA_BLOCK "Alarm_Axis_Position_Function_Infeed"   // DB43
{ S7_Optimized_Access := 'FALSE' }
VERSION : 0.1
// stored: InstanceOfName Alarm_Axis_Position_Function
"Alarm_Axis_Position_Function"
BEGIN
END_DATA_BLOCK

DATA_BLOCK "DriveConfirmation_Function_Axis1"   // DB45
{ S7_Optimized_Access := 'FALSE' }
VERSION : 0.1
// stored: InstanceOfName DriveConfirmation_Function
"DriveConfirmation_Function"
BEGIN
END_DATA_BLOCK

DATA_BLOCK "DriveConfirmation_Function_Axis2"   // DB46
{ S7_Optimized_Access := 'FALSE' }
VERSION : 0.1
// stored: InstanceOfName DriveConfirmation_Function
"DriveConfirmation_Function"
BEGIN
END_DATA_BLOCK

DATA_BLOCK "DriveConfirmation_Function_Axis 3"   // DB47
{ S7_Optimized_Access := 'FALSE' }
VERSION : 0.1
// stored: InstanceOfName DriveConfirmation_Function
"DriveConfirmation_Function"
BEGIN
END_DATA_BLOCK

DATA_BLOCK "DriveConfirmation_Function_Axis 4"   // DB48
{ S7_Optimized_Access := 'FALSE' }
VERSION : 0.1
// stored: InstanceOfName DriveConfirmation_Function
"DriveConfirmation_Function"
BEGIN
END_DATA_BLOCK

DATA_BLOCK "DriveConfirmation_Function_Axis 5"   // DB49
{ S7_Optimized_Access := 'FALSE' }
VERSION : 0.1
// stored: InstanceOfName DriveConfirmation_Function
"DriveConfirmation_Function"
BEGIN
END_DATA_BLOCK

// folder: Motion

DATA_BLOCK "PositionManagement"   // DB51
{ S7_Optimized_Access := 'FALSE' }
VERSION : 0.1
   VAR
      Data : Struct   // Data
         CntPlsPrev : DInt := 0;   // Flowpulsen vorige scan
         CntPlsDiff : DInt := 0;   // Flowpulsen verschil
         CntPlsAct : DInt := 0;   // Flowpulsen actueel
         DosActueel : Real := 0.0;   // Dosering actueel ('x' gram/liter/kg gist)
         Actual_Axis3_Position : Real;   // Actual Position of Axis 3 stored in this datablock
         Actual_Axis1_Position : Real;
      END_STRUCT;
      "Axis 3" : Struct
         Values : Struct
            AxisName : String := 'Drive 3 - Wals';
            "Reference Position" : Int := 0;
            "Set Position" : Real := -50.0;
            "Rest Position" : Real := -25.0;
            Acceleration : Real := 0.0;
            Deacceleration : Real;
            "Axis Correction" : Real := 1.0E-06;
            "Position Offset" : Real := 35.0;
            Pulsfactor : Real := 0.82;
            Axis_Speed : Int := 0;
         END_STRUCT;
         Commands : Struct
            "Go To Rest" : Bool;
            "Start Ref Run" : Bool;
            "Take Over Pos" : Bool;
            "Go To Position" : Bool;
            "Jog Fwd" : Bool;
            "Jog Rev" : Bool;
            Axis_Brake : Bool;
            MasterWord : String;
            "Master Callback" : String;
         END_STRUCT;
         Messages : Struct
            "Axis Busy" : Bool;
            "Error Executing Command" : Bool;
            "Axis On Rest" : Bool;
            "Axis On Position" : Bool;
            "Drive State (Option)" : String;
            "Slip State" : String;
            AxisHasReference : Bool;
         END_STRUCT;
      END_STRUCT;
      Demo_Pos : Struct
         Desired_Pos : Real;
         Start : Bool;
         SetRefRunActive : Bool;
         RequestMove1 : Bool;
         RequestMove2 : Bool;
         PositionMove2 : Real := -330.0;
         PositionMove1 : Real := -120.0;
         Pos2Done : Bool;
         BrakeOnPos1 : Bool;
         BrakeOnPos2 : Bool;
         ManualSensorOverride : Bool;
      END_STRUCT;
      Axis_1 : Struct
         Values : Struct
            AxisName : String := 'Drive 1 - Infeed';
            "Reference Position" : Int := 0;
            "Set Position" : Real := 0.0;
            "Rest Position" : Real := 0.0;
            Acceleration : Real := 0.0;
            Deacceleration : Real;
            "Axis Correction" : Real := 1.0E-06;
            "Position Offset" : Real := 0.001;
            Pulsfactor : Real := -0.325;
            Axis_Speed : Int := 0;
         END_STRUCT;
         Commands : Struct
            "Go To Rest" : Bool;
            "Start Ref Run" : Bool;
            "Take Over Pos" : Bool;
            "Go To Position" : Bool;
            "Jog Fwd" : Bool;
            "Jog Rev" : Bool;
            Axis_Brake : Bool;
            ReferenceSwitch : Bool;
            MasterWord : String;
            "Master Callback" : String;
         END_STRUCT;
         Messages : Struct
            "Axis Busy" : Bool;
            "Error Executing Command" : Bool;
            "Axis On Rest" : Bool;
            "Axis On Position" : Bool;
            "Drive State (Option)" : String;
            "Slip State" : String;
            AxisHasReference : Bool;
         END_STRUCT;
      END_STRUCT;
   END_VAR
BEGIN
END_DATA_BLOCK

DATA_BLOCK "MC_Move_Prog.1"   // DB54
{ S7_Optimized_Access := 'FALSE' }
VERSION : 0.1
// stored: InstanceOfName MC_Move
"MC_Move"
BEGIN
END_DATA_BLOCK

DATA_BLOCK "MC_Jog_OB1"   // DB56
{ S7_Optimized_Access := 'FALSE' }
VERSION : 0.1
// stored: InstanceOfName MC_Jog
"MC_Jog"
BEGIN
END_DATA_BLOCK

DATA_BLOCK "EncoderFeedback_Band"   // DB89
{ S7_Optimized_Access := 'FALSE' }
VERSION : 0.1
// stored: InstanceOfName FB_EncoderFeedback_Lineair
"FB_EncoderFeedback_Lineair"
BEGIN
END_DATA_BLOCK

// folder: (top level)

FUNCTION "3 - Prog. 1" : Void   // FC1, LAD
TITLE = System Program 1
{ S7_Optimized_Access := 'FALSE' }
VERSION : 0.1
// DF
   VAR_INPUT
      Axis_3_MovePosition1 : Real;
      Axis_3_MovePosition2 : Real;
   END_VAR
   VAR_OUTPUT
      Axis_On_Pos_1 : Bool;
      Axis_On_Pos_2 : Bool;
   END_VAR
   VAR_TEMP
      TempProdCounter : Int;
      Temp_ProductsToProduce : Bool;
      TimerRunning : Bool;
      ProduceContact : Bool;
      Move2Done : Bool;
      SRWals : Bool;
      Move2Busy : Bool;
      SR_Move2 : Bool;
      Move1Busy : Bool;
      P_TRIG_SnrBand : Bool;
      Temp1 : Bool;
      Min_Pos_1 : Real;
      Max_Pos_1 : Real;
      Min_Pos_2 : Real;
      Max_Pos_2 : Real;
      SR_Move3 : Bool;
      SR_Move1 : Bool;
      AxisToRest : Bool;
      SubDone : Bool;
      P_Trig_ProBehWals : Bool;
      ProductsBehindWals : Int;
      ProductBehindWals : Bool;
      AandrukCilindersOut : Bool;
      Retourband_Delayed : Bool;
      BlowOff_Activated : Bool;
      Pos2_Done : Bool;
      Pos1_Done : Bool;
      ToWaitPosition : Bool;
      BlowOffConf : Bool;
      PTrig_Blow : Bool;
      Move2Done_2 : Bool;
      GoToMove2Pos : Bool;
   END_VAR
   VAR_TEMP   // added for the SCL form of the ladder/FBD networks
      _w1 : Bool;
   END_VAR
BEGIN

REGION Network 1: Set Counter on Zero
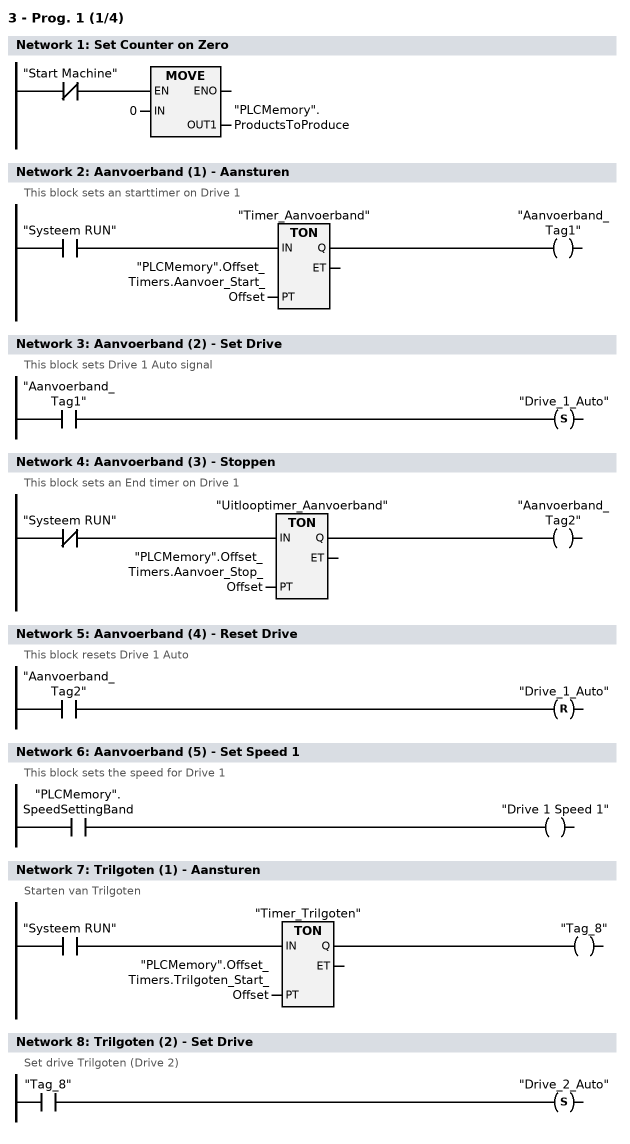
   RUNG wire#powerrail
      I_Contact( "Start Machine" )
      { S7_GenerateENO := "TRUE" } Move(in := 0, out1 => "PLCMemory".ProductsToProduce)
   END_RUNG
   // the same network as SCL:
   IF NOT "Start Machine" THEN "PLCMemory".ProductsToProduce := 0; END_IF;
END_REGION

REGION Network 2: Aanvoerband (1) - Aansturen
   // This block sets an starttimer on Drive 1
   "Timer_Aanvoerband".TON(IN := "Systeem RUN", PT := "PLCMemory".Offset_Timers.Aanvoer_Start_Offset);
   "Aanvoerband_Tag1" := "Timer_Aanvoerband".Q;
END_REGION

REGION Network 3: Aanvoerband (2) - Set Drive
   // This block sets Drive 1 Auto signal
   RUNG wire#powerrail
      Contact( "Aanvoerband_Tag1" )
      S_Coil( "Drive_1_Auto" )
   END_RUNG
   // the same network as SCL:
   IF "Aanvoerband_Tag1" THEN "Drive_1_Auto" := TRUE; END_IF;
END_REGION

REGION Network 4: Aanvoerband (3) - Stoppen
   // This block sets an End timer on Drive 1
   "Uitlooptimer_Aanvoerband".TON(IN := NOT "Systeem RUN", PT := "PLCMemory".Offset_Timers.Aanvoer_Stop_Offset);
   "Aanvoerband_Tag2" := "Uitlooptimer_Aanvoerband".Q;
END_REGION

REGION Network 5: Aanvoerband (4) - Reset Drive
   // This block resets Drive 1 Auto
   RUNG wire#powerrail
      Contact( "Aanvoerband_Tag2" )
      R_Coil( "Drive_1_Auto" )
   END_RUNG
   // the same network as SCL:
   IF "Aanvoerband_Tag2" THEN "Drive_1_Auto" := FALSE; END_IF;
END_REGION

REGION Network 6: Aanvoerband (5) - Set Speed 1
   // This block sets the speed for Drive 1
   RUNG wire#powerrail
      Contact( "PLCMemory".SpeedSettingBand )
      Coil( "Drive 1 Speed 1" )
   END_RUNG
   // the same network as SCL:
   "Drive 1 Speed 1" := "PLCMemory".SpeedSettingBand;
END_REGION

REGION Network 7: Trilgoten (1) - Aansturen
   // Starten van Trilgoten
   "Timer_Trilgoten".TON(IN := "Systeem RUN", PT := "PLCMemory".Offset_Timers.Trilgoten_Start_Offset);
   "Tag_8" := "Timer_Trilgoten".Q;
END_REGION

REGION Network 8: Trilgoten (2) - Set Drive
   // Set drive Trilgoten (Drive 2)
   RUNG wire#powerrail
      Contact( "Tag_8" )
      S_Coil( "Drive_2_Auto" )
   END_RUNG
   // the same network as SCL:
   IF "Tag_8" THEN "Drive_2_Auto" := TRUE; END_IF;
END_REGION

REGION Network 9: Trilgoten (3) - Stoppen
   // Stoppen van de trilgoten.
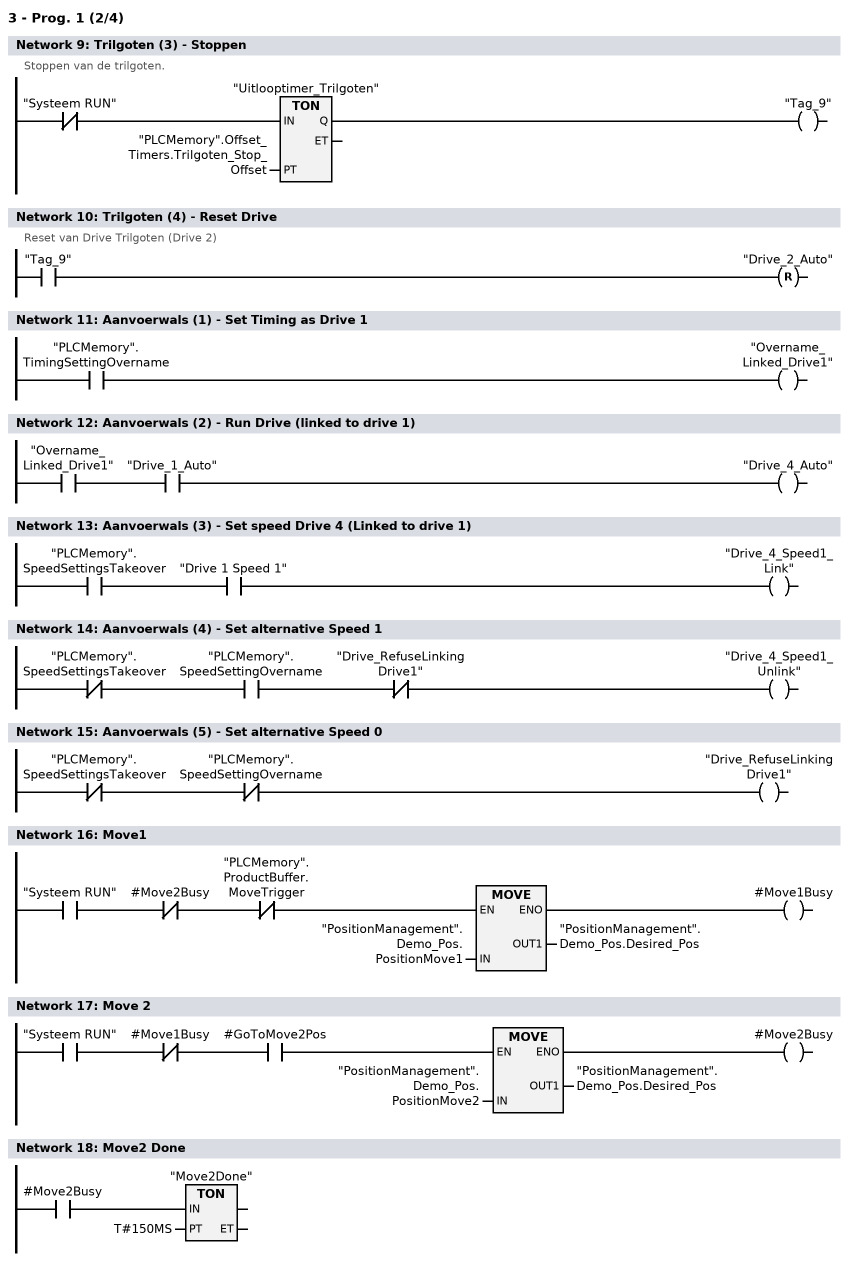
   "Uitlooptimer_Trilgoten".TON(IN := NOT "Systeem RUN", PT := "PLCMemory".Offset_Timers.Trilgoten_Stop_Offset);
   "Tag_9" := "Uitlooptimer_Trilgoten".Q;
END_REGION

REGION Network 10: Trilgoten (4) - Reset Drive
   // Reset van Drive Trilgoten (Drive 2)
   RUNG wire#powerrail
      Contact( "Tag_9" )
      R_Coil( "Drive_2_Auto" )
   END_RUNG
   // the same network as SCL:
   IF "Tag_9" THEN "Drive_2_Auto" := FALSE; END_IF;
END_REGION

REGION Network 11: Aanvoerwals (1) - Set Timing as Drive 1
   RUNG wire#powerrail
      Contact( "PLCMemory".TimingSettingOvername )
      Coil( "Overname_Linked_Drive1" )
   END_RUNG
   // the same network as SCL:
   "Overname_Linked_Drive1" := "PLCMemory".TimingSettingOvername;
END_REGION

REGION Network 12: Aanvoerwals (2) - Run Drive (linked to drive 1)
   RUNG wire#powerrail
      Contact( "Overname_Linked_Drive1" )
      Contact( "Drive_1_Auto" )
      Coil( "Drive_4_Auto" )
   END_RUNG
   // the same network as SCL:
   "Drive_4_Auto" := "Overname_Linked_Drive1" AND "Drive_1_Auto";
END_REGION

REGION Network 13: Aanvoerwals (3) - Set speed Drive 4 (Linked to drive 1)
   RUNG wire#powerrail
      Contact( "PLCMemory".SpeedSettingsTakeover )
      Contact( "Drive 1 Speed 1" )
      Coil( "Drive_4_Speed1_Link" )
   END_RUNG
   // the same network as SCL:
   "Drive_4_Speed1_Link" := "PLCMemory".SpeedSettingsTakeover AND "Drive 1 Speed 1";
END_REGION

REGION Network 14: Aanvoerwals (4) - Set alternative Speed 1
   RUNG wire#powerrail
      I_Contact( "PLCMemory".SpeedSettingsTakeover )
      Contact( "PLCMemory".SpeedSettingOvername )
      I_Contact( "Drive_RefuseLinkingDrive1" )
      Coil( "Drive_4_Speed1_Unlink" )
   END_RUNG
   // the same network as SCL:
   "Drive_4_Speed1_Unlink" := NOT "PLCMemory".SpeedSettingsTakeover AND "PLCMemory".SpeedSettingOvername AND NOT "Drive_RefuseLinkingDrive1";
END_REGION

REGION Network 15: Aanvoerwals (5) - Set alternative Speed 0
   RUNG wire#powerrail
      I_Contact( "PLCMemory".SpeedSettingsTakeover )
      I_Contact( "PLCMemory".SpeedSettingOvername )
      Coil( "Drive_RefuseLinkingDrive1" )
   END_RUNG
   // the same network as SCL:
   "Drive_RefuseLinkingDrive1" := NOT "PLCMemory".SpeedSettingsTakeover AND NOT "PLCMemory".SpeedSettingOvername;
END_REGION

REGION Network 16: Move1
   RUNG wire#powerrail
      Contact( "Systeem RUN" )
      I_Contact( #Move2Busy )
      I_Contact( "PLCMemory".ProductBuffer.MoveTrigger )
      { S7_GenerateENO := "TRUE" } Move(in := "PositionManagement".Demo_Pos.PositionMove1, out1 => "PositionManagement".Demo_Pos.Desired_Pos)
      Coil( #Move1Busy )
   END_RUNG
   // the same network as SCL:
   // ENO of a box is taken as its EN; it also drops when the box reports an error
   #_w1 := "Systeem RUN" AND NOT #Move2Busy AND NOT "PLCMemory".ProductBuffer.MoveTrigger;
   IF #_w1 THEN
       "PositionManagement".Demo_Pos.Desired_Pos := "PositionManagement".Demo_Pos.PositionMove1;
   END_IF;
   #Move1Busy := #_w1;
END_REGION

REGION Network 17: Move 2
   RUNG wire#powerrail
      Contact( "Systeem RUN" )
      I_Contact( #Move1Busy )
      Contact( #GoToMove2Pos )
      { S7_GenerateENO := "TRUE" } Move(in := "PositionManagement".Demo_Pos.PositionMove2, out1 => "PositionManagement".Demo_Pos.Desired_Pos)
      Coil( #Move2Busy )
   END_RUNG
   // the same network as SCL:
   // ENO of a box is taken as its EN; it also drops when the box reports an error
   #_w1 := "Systeem RUN" AND NOT #Move1Busy AND #GoToMove2Pos;
   IF #_w1 THEN
       "PositionManagement".Demo_Pos.Desired_Pos := "PositionManagement".Demo_Pos.PositionMove2;
   END_IF;
   #Move2Busy := #_w1;
END_REGION

REGION Network 18: Move2 Done
   "Move2Done".TON(IN := #Move2Busy, PT := T#150MS);
END_REGION

REGION Network 19: Set Move 2